   "20_TANKS_IP_DATA_RIO_04_FIRST_TANK_BWT_TEMP" : Real = PLC "20_TANKS_IP_DATA".RIO_04.FIRST_TANK.BWT_TEMP, 1 s
   "20_TANKS_IP_DATA_RIO_04_FIRST_TANK_BWT_DO" : Real = PLC "20_TANKS_IP_DATA".RIO_04.FIRST_TANK.BWT_DO, 1 s
   "20_TANKS_IP_DATA_RIO_04_FIRST_TANK_BWT_PH" : Real = PLC "20_TANKS_IP_DATA".RIO_04.FIRST_TANK.BWT_PH, 1 s
   "20_TANKS_IP_DATA_RIO_06_FIRST_TANK_BWT_TEMP" : Real = PLC "20_TANKS_IP_DATA".RIO_06.FIRST_TANK.BWT_TEMP, 1 s
   "20_TANKS_IP_DATA_RIO_04_FIRST_TANK_BWT_LEVEL" : Real = PLC "20_TANKS_IP_DATA".RIO_04.FIRST_TANK.BWT_LEVEL, 1 s
   "504_Tank Grouping_DB2020_Tank12 Min Time_ET" : Time = PLC "504_Tank Grouping_DB2020"."Tank12 Min Time".ET, 1 s
   "20_TANKS_IP_DATA_RIO_06_SECOND_TANK_BWT_LEVEL" : Real = PLC "20_TANKS_IP_DATA".RIO_06.SECOND_TANK.BWT_LEVEL, 1 s
   "504_Tank Grouping_DB2020_Time Left Tank_Time Left Tank 13" : Real = PLC "504_Tank Grouping_DB2020"."Time Left Tank"."Time Left Tank 13", 1 s
   "504_Tank Grouping_DB2020_Time Left Tank_Time Left Tank 12" : Real = PLC "504_Tank Grouping_DB2020"."Time Left Tank"."Time Left Tank 12", 1 s
   "504_Tank Grouping_DB2020_Time Left Tank_Time Left Tank 11" : Real = PLC "504_Tank Grouping_DB2020"."Time Left Tank"."Time Left Tank 11", 1 s
   "504_Tank Grouping_DB2020_Time Left Tank_Time Left Tank 10" : Real = PLC "504_Tank Grouping_DB2020"."Time Left Tank"."Time Left Tank 10", 1 s
   "504_Tank Grouping_DB2020_Time Left Tank_Time Left Tank 9" : Real = PLC "504_Tank Grouping_DB2020"."Time Left Tank"."Time Left Tank 9", 1 s
   "504_Tank Grouping_DB2020_Time Left Tank_Time Left Tank 8" : Real = PLC "504_Tank Grouping_DB2020"."Time Left Tank"."Time Left Tank 8", 1 s
   "504_Tank Grouping_DB2020_Time Left Tank_Time Left Tank 6" : Real = PLC "504_Tank Grouping_DB2020"."Time Left Tank"."Time Left Tank 6", 1 s
   "504_Tank Grouping_DB2020_Time Left Tank_Time Left Tank 5" : Real = PLC "504_Tank Grouping_DB2020"."Time Left Tank"."Time Left Tank 5", 1 s
   "504_Tank Grouping_DB2020_Time Left Tank_Time Left Tank 4" : Real = PLC "504_Tank Grouping_DB2020"."Time Left Tank"."Time Left Tank 4", 1 s
   "504_Tank Grouping_DB2020_Time Left Tank_Time Left Tank 3" : Real = PLC "504_Tank Grouping_DB2020"."Time Left Tank"."Time Left Tank 3", 1 s
   "504_Tank Grouping_DB2020_Time Left Tank_Time Left Tank 2" : Real = PLC "504_Tank Grouping_DB2020"."Time Left Tank"."Time Left Tank 2", 1 s
   "504_Tank Grouping_DB2020_Time Left Tank_Time Left Tank 7" : Real = PLC "504_Tank Grouping_DB2020"."Time Left Tank"."Time Left Tank 7", 1 s
   "504_Tank Grouping_DB2020_Offset Timer_ET" : Time = PLC "504_Tank Grouping_DB2020"."Offset Timer".ET, 1 s
   "80_From_HMI_Test Tank Request" : Bool = PLC "80_From_HMI"."Test Tank Request", 1 s
   "504_Tank Grouping_DB2020_RUN" : Bool = PLC "504_Tank Grouping_DB2020".RUN, 1 s
   "20_TANKS_IP_DATA_RIO_07_FIRST_TANK_BWT_TEMP" : Real = PLC "20_TANKS_IP_DATA".RIO_07.FIRST_TANK.BWT_TEMP, 1 s
   "20_TANKS_IP_DATA_RIO_07_FIRST_TANK_BWT_DO" : Real = PLC "20_TANKS_IP_DATA".RIO_07.FIRST_TANK.BWT_DO, 1 s
   "20_TANKS_IP_DATA_RIO_07_FIRST_TANK_BWT_PH" : Real = PLC "20_TANKS_IP_DATA".RIO_07.FIRST_TANK.BWT_PH, 1 s
   "20_TANKS_IP_DATA_RIO_07_FIRST_TANK_BWT_LEVEL" : Real = PLC "20_TANKS_IP_DATA".RIO_07.FIRST_TANK.BWT_LEVEL, 1 s
   "20_TANKS_IP_DATA_RIO_07_FIRST_TANK_TANKS_PRESS" : Real = PLC "20_TANKS_IP_DATA".RIO_07.FIRST_TANK.TANKS_PRESS, 1 s
   "504_Tank Grouping_DB2020_Tank14 Min Time_ET" : Time = PLC "504_Tank Grouping_DB2020"."Tank14 Min Time".ET, 1 s
   "504_Tank Grouping_DB2020_Tank13 Min Time_ET" : Time = PLC "504_Tank Grouping_DB2020"."Tank13 Min Time".ET, 1 s
   "20_TANKS_IP_DATA_RIO_06_SECOND_TANK_BWT_TEMP" : Real = PLC "20_TANKS_IP_DATA".RIO_06.SECOND_TANK.BWT_TEMP, 1 s
   "20_TANKS_IP_DATA_RIO_06_SECOND_TANK_BWT_DO" : Real = PLC "20_TANKS_IP_DATA".RIO_06.SECOND_TANK.BWT_DO, 1 s
   "20_TANKS_IP_DATA_RIO_06_SECOND_TANK_BWT_PH" : Real = PLC "20_TANKS_IP_DATA".RIO_06.SECOND_TANK.BWT_PH, 1 s
   "20_TANKS_IP_DATA_RIO_06_SECOND_TANK_TANKS_PRESS" : Real = PLC "20_TANKS_IP_DATA".RIO_06.SECOND_TANK.TANKS_PRESS, 1 s
   "20_TANKS_IP_DATA_RIO_04_FIRST_TANK_TANKS_PRESS" : Real = PLC "20_TANKS_IP_DATA".RIO_04.FIRST_TANK.TANKS_PRESS, 1 s
   "504_Tank Grouping_DB2020_Tank7 Min Time_ET" : Time = PLC "504_Tank Grouping_DB2020"."Tank7 Min Time".ET, 1 s
   "20_TANKS_IP_DATA_RIO_03_SECOND_TANK_BWT_TEMP" : Real = PLC "20_TANKS_IP_DATA".RIO_03.SECOND_TANK.BWT_TEMP, 1 s
   "504_Tank Grouping_DB2020_Sequence Time m Offset" : Time = PLC "504_Tank Grouping_DB2020"."Sequence Time m Offset", 1 s
   "504_Tank Grouping_DB2020_RUN TANK 13" : Bool = PLC "504_Tank Grouping_DB2020"."RUN TANK 13", 1 s
   "504_Tank Grouping_DB2020_RUN TANK 12" : Bool = PLC "504_Tank Grouping_DB2020"."RUN TANK 12", 1 s
   "504_Tank Grouping_DB2020_RUN TANK 11" : Bool = PLC "504_Tank Grouping_DB2020"."RUN TANK 11", 1 s
   "504_Tank Grouping_DB2020_RUN TANK 10" : Bool = PLC "504_Tank Grouping_DB2020"."RUN TANK 10", 1 s
   "504_Tank Grouping_DB2020_RUN TANK 9" : Bool = PLC "504_Tank Grouping_DB2020"."RUN TANK 9", 1 s
   "504_Tank Grouping_DB2020_RUN TANK 8" : Bool = PLC "504_Tank Grouping_DB2020"."RUN TANK 8", 1 s
   "504_Tank Grouping_DB2020_RUN TANK 6" : Bool = PLC "504_Tank Grouping_DB2020"."RUN TANK 6", 1 s
   "504_Tank Grouping_DB2020_RUN TANK 14" : Bool = PLC "504_Tank Grouping_DB2020"."RUN TANK 14", 1 s
   "20_TANKS_IP_DATA_RIO_07_FIRST_TANK_MBG_FLOW" : Real = PLC "20_TANKS_IP_DATA".RIO_07.FIRST_TANK.MBG_FLOW, 1 s
   "20_TANKS_IP_DATA_RIO_07_FIRST_TANK_USD_FLOW" : Real = PLC "20_TANKS_IP_DATA".RIO_07.FIRST_TANK.USD_FLOW, 1 s
   "20_TANKS_IP_DATA_RIO_07_FIRST_TANK_GTT_ISOL_VALVE_CLSD" : Bool = PLC "20_TANKS_IP_DATA".RIO_07.FIRST_TANK.GTT_ISOL_VALVE_CLSD, 1 s
   "20_TANKS_IP_DATA_RIO_07_FIRST_TANK_GTT_ISOL_VALVE_OPEN" : Bool = PLC "20_TANKS_IP_DATA".RIO_07.FIRST_TANK.GTT_ISOL_VALVE_OPEN, 1 s
   "20_TANKS_IP_DATA_RIO_07_FIRST_TANK_BWT_LEVEL_HIHI" : Bool = PLC "20_TANKS_IP_DATA".RIO_07.FIRST_TANK.BWT_LEVEL_HIHI, 1 s
   "20_TANKS_IP_DATA_RIO_06_SECOND_TANK_GTT_ISOL_VALVE_CLSD" : Bool = PLC "20_TANKS_IP_DATA".RIO_06.SECOND_TANK.GTT_ISOL_VALVE_CLSD, 1 s
   "20_TANKS_IP_DATA_RIO_06_SECOND_TANK_GTT_ISOL_VALVE_OPEN" : Bool = PLC "20_TANKS_IP_DATA".RIO_06.SECOND_TANK.GTT_ISOL_VALVE_OPEN, 1 s
   "Tank 3S BWT Level High High Switch" : Bool = PLC "Tank 3S BWT Level High High Switch" AT %I33.2, 1 s
   "20_TANKS_IP_DATA_RIO_06_SECOND_TANK_USD_FLOW" : Real = PLC "20_TANKS_IP_DATA".RIO_06.SECOND_TANK.USD_FLOW, 1 s
   "20_TANKS_IP_DATA_RIO_06_SECOND_TANK_BWT_LEVEL_HIHI" : Bool = PLC "20_TANKS_IP_DATA".RIO_06.SECOND_TANK.BWT_LEVEL_HIHI, 1 s
   "20_TANKS_IP_DATA_RIO_06_FIRST_TANK_GTT_ISOL_VALVE_CLSD" : Bool = PLC "20_TANKS_IP_DATA".RIO_06.FIRST_TANK.GTT_ISOL_VALVE_CLSD, 1 s
   "20_TANKS_IP_DATA_RIO_06_FIRST_TANK_GTT_ISOL_VALVE_OPEN" : Bool = PLC "20_TANKS_IP_DATA".RIO_06.FIRST_TANK.GTT_ISOL_VALVE_OPEN, 1 s
   "20_TANKS_IP_DATA_RIO_06_FIRST_TANK_MBG_FLOW" : Real = PLC "20_TANKS_IP_DATA".RIO_06.FIRST_TANK.MBG_FLOW, 1 s
   "20_TANKS_IP_DATA_RIO_06_FIRST_TANK_USD_FLOW" : Real = PLC "20_TANKS_IP_DATA".RIO_06.FIRST_TANK.USD_FLOW, 1 s
   "20_TANKS_IP_DATA_RIO_06_FIRST_TANK_BWT_LEVEL_HIHI" : Bool = PLC "20_TANKS_IP_DATA".RIO_06.FIRST_TANK.BWT_LEVEL_HIHI, 1 s
   "20_TANKS_IP_DATA_RIO_05_SECOND_TANK_GTT_ISOL_VALVE_CLSD" : Bool = PLC "20_TANKS_IP_DATA".RIO_05.SECOND_TANK.GTT_ISOL_VALVE_CLSD, 1 s
   "20_TANKS_IP_DATA_RIO_01_FIRST_TANK_TANKS_PRESS" : Real = PLC "20_TANKS_IP_DATA".RIO_01.FIRST_TANK.TANKS_PRESS, 1 s
   "20_TANKS_IP_DATA_RIO_01_FIRST_TANK_BWT_LEVEL" : Real = PLC "20_TANKS_IP_DATA".RIO_01.FIRST_TANK.BWT_LEVEL, 1 s
   "20_TANKS_IP_DATA_RIO_01_FIRST_TANK_BWT_PH" : Real = PLC "20_TANKS_IP_DATA".RIO_01.FIRST_TANK.BWT_PH, 1 s
   "20_TANKS_IP_DATA_RIO_01_FIRST_TANK_BWT_DO" : Real = PLC "20_TANKS_IP_DATA".RIO_01.FIRST_TANK.BWT_DO, 1 s
   "20_TANKS_IP_DATA_RIO_03_SECOND_TANK_BWT_DO" : Real = PLC "20_TANKS_IP_DATA".RIO_03.SECOND_TANK.BWT_DO, 1 s
   "20_TANKS_IP_DATA_RIO_03_SECOND_TANK_BWT_PH" : Real = PLC "20_TANKS_IP_DATA".RIO_03.SECOND_TANK.BWT_PH, 1 s
   "20_TANKS_IP_DATA_RIO_03_SECOND_TANK_BWT_LEVEL" : Real = PLC "20_TANKS_IP_DATA".RIO_03.SECOND_TANK.BWT_LEVEL, 1 s
   "20_TANKS_IP_DATA_RIO_03_SECOND_TANK_TANKS_PRESS" : Real = PLC "20_TANKS_IP_DATA".RIO_03.SECOND_TANK.TANKS_PRESS, 1 s
   "504_Tank Grouping_DB2020_Tank6 Min Time_ET" : Time = PLC "504_Tank Grouping_DB2020"."Tank6 Min Time".ET, 1 s
   "20_TANKS_IP_DATA_RIO_03_FIRST_TANK_BWT_TEMP" : Real = PLC "20_TANKS_IP_DATA".RIO_03.FIRST_TANK.BWT_TEMP, 1 s
   "20_TANKS_IP_DATA_RIO_03_FIRST_TANK_BWT_DO" : Real = PLC "20_TANKS_IP_DATA".RIO_03.FIRST_TANK.BWT_DO, 1 s
   "20_TANKS_IP_DATA_RIO_03_FIRST_TANK_BWT_PH" : Real = PLC "20_TANKS_IP_DATA".RIO_03.FIRST_TANK.BWT_PH, 1 s
   "20_TANKS_IP_DATA_RIO_03_FIRST_TANK_BWT_LEVEL" : Real = PLC "20_TANKS_IP_DATA".RIO_03.FIRST_TANK.BWT_LEVEL, 1 s
   "20_TANKS_IP_DATA_RIO_03_FIRST_TANK_TANKS_PRESS" : Real = PLC "20_TANKS_IP_DATA".RIO_03.FIRST_TANK.TANKS_PRESS, 1 s
   "504_Tank Grouping_DB2020_Tank5 Min Time_ET" : Time = PLC "504_Tank Grouping_DB2020"."Tank5 Min Time".ET, 1 s
   "504_Tank Grouping_DB2020_Tank3 Min Time_ET" : Time = PLC "504_Tank Grouping_DB2020"."Tank3 Min Time".ET, 1 s
   "20_TANKS_IP_DATA_RIO_05_SECOND_TANK_MBG_FLOW" : Real = PLC "20_TANKS_IP_DATA".RIO_05.SECOND_TANK.MBG_FLOW, 1 s
   "504_Tank Grouping_DB2020_Tank4 Min Time_ET" : Time = PLC "504_Tank Grouping_DB2020"."Tank4 Min Time".ET, 1 s
   "20_TANKS_IP_DATA_RIO_01_THIRD_TANK_BWT_DO" : Real = PLC "20_TANKS_IP_DATA".RIO_01.THIRD_TANK.BWT_DO, 1 s
   "20_TANKS_IP_DATA_RIO_01_THIRD_TANK_BWT_PH" : Real = PLC "20_TANKS_IP_DATA".RIO_01.THIRD_TANK.BWT_PH, 1 s
   "20_TANKS_IP_DATA_RIO_01_THIRD_TANK_BWT_LEVEL" : Real = PLC "20_TANKS_IP_DATA".RIO_01.THIRD_TANK.BWT_LEVEL, 1 s
   "20_TANKS_IP_DATA_RIO_01_THIRD_TANK_TANKS_PRESS" : Real = PLC "20_TANKS_IP_DATA".RIO_01.THIRD_TANK.TANKS_PRESS, 1 s
   "20_TANKS_IP_DATA_RIO_01_SECOND_TANK_BWT_TEMP" : Real = PLC "20_TANKS_IP_DATA".RIO_01.SECOND_TANK.BWT_TEMP, 1 s
   "20_TANKS_IP_DATA_RIO_01_SECOND_TANK_BWT_DO" : Real = PLC "20_TANKS_IP_DATA".RIO_01.SECOND_TANK.BWT_DO, 1 s
   "20_TANKS_IP_DATA_RIO_01_SECOND_TANK_BWT_PH" : Real = PLC "20_TANKS_IP_DATA".RIO_01.SECOND_TANK.BWT_PH, 1 s
   "20_TANKS_IP_DATA_RIO_01_SECOND_TANK_BWT_LEVEL" : Real = PLC "20_TANKS_IP_DATA".RIO_01.SECOND_TANK.BWT_LEVEL, 1 s
   "20_TANKS_IP_DATA_RIO_01_SECOND_TANK_TANKS_PRESS" : Real = PLC "20_TANKS_IP_DATA".RIO_01.SECOND_TANK.TANKS_PRESS, 1 s
   "504_Tank Grouping_DB2020_Tank2 Min Time_ET" : Time = PLC "504_Tank Grouping_DB2020"."Tank2 Min Time".ET, 1 s
   "504_Tank Grouping_DB2020_Tank1 Min Time_ET" : Time = PLC "504_Tank Grouping_DB2020"."Tank1 Min Time".ET, 1 s
   "20_TANKS_IP_DATA_RIO_01_FIRST_TANK_BWT_TEMP" : Real = PLC "20_TANKS_IP_DATA".RIO_01.FIRST_TANK.BWT_TEMP, 1 s
   "20_TANKS_IP_DATA_RIO_01_THIRD_TANK_BWT_TEMP" : Real = PLC "20_TANKS_IP_DATA".RIO_01.THIRD_TANK.BWT_TEMP, 1 s
   "RIO3_SPR_DI_33_3" : Bool = PLC RIO3_SPR_DI_33_3 AT %I33.3, 1 s
   "150_GCU_LCL_CNTRL_DB_LCL_CNTRL_ACTV" : Bool = PLC "150_GCU_LCL_CNTRL_DB".LCL_CNTRL_ACTV, 1 s
   "RIO3_SPR_DI_33_5" : Bool = PLC RIO3_SPR_DI_33_5 AT %I33.5, 1 s
   "TT426_5S_ALM_ANALOG_DB_VERY LOW LEVEL VALUE (LL)" : Real = PLC TT426_5S_ALM_ANALOG_DB."VERY LOW LEVEL VALUE (LL)" AT %DB2082.DBD22, 1 s
   "TT426_5S_ALM_ANALOG_DB_LOW LEVEL VALUE (L)" : Real = PLC TT426_5S_ALM_ANALOG_DB."LOW LEVEL VALUE (L)" AT %DB2082.DBD26, 1 s
   "TT426_5S_ALM_ANALOG_DB_HIGH LEVEL VALUE (H)" : Real = PLC TT426_5S_ALM_ANALOG_DB."HIGH LEVEL VALUE (H)" AT %DB2082.DBD30, 1 s
   "TT426_5S_ALM_ANALOG_DB_VERY HIGH LEVEL VALUE (HH)" : Real = PLC TT426_5S_ALM_ANALOG_DB."VERY HIGH LEVEL VALUE (HH)" AT %DB2082.DBD34, 1 s
   "TT426STR_ALM_ANALOG_DB_VERY LOW LEVEL VALUE (LL)" : Real = PLC TT426STR_ALM_ANALOG_DB."VERY LOW LEVEL VALUE (LL)" AT %DB2072.DBD22, 1 s
   "TT426STR_ALM_ANALOG_DB_LOW LEVEL VALUE (L)" : Real = PLC TT426STR_ALM_ANALOG_DB."LOW LEVEL VALUE (L)" AT %DB2072.DBD26, 1 s
   "TT426STR_ALM_ANALOG_DB_HIGH LEVEL VALUE (H)" : Real = PLC TT426STR_ALM_ANALOG_DB."HIGH LEVEL VALUE (H)" AT %DB2072.DBD30, 1 s
   "TT426STR_ALM_ANALOG_DB_VERY HIGH LEVEL VALUE (HH)" : Real = PLC TT426STR_ALM_ANALOG_DB."VERY HIGH LEVEL VALUE (HH)" AT %DB2072.DBD34, 1 s
   "TT426PORT_ALM_ANALOG_DB_VERY LOW LEVEL VALUE (LL)" : Real = PLC TT426PORT_ALM_ANALOG_DB."VERY LOW LEVEL VALUE (LL)" AT %DB2071.DBD22, 1 s
   "TT426PORT_ALM_ANALOG_DB_LOW LEVEL VALUE (L)" : Real = PLC TT426PORT_ALM_ANALOG_DB."LOW LEVEL VALUE (L)" AT %DB2071.DBD26, 1 s
   "TT426PORT_ALM_ANALOG_DB_HIGH LEVEL VALUE (H)" : Real = PLC TT426PORT_ALM_ANALOG_DB."HIGH LEVEL VALUE (H)" AT %DB2071.DBD30, 1 s
   "TT426PORT_ALM_ANALOG_DB_VERY HIGH LEVEL VALUE (HH)" : Real = PLC TT426PORT_ALM_ANALOG_DB."VERY HIGH LEVEL VALUE (HH)" AT %DB2071.DBD34, 1 s
   "PIT424PORT_ALM_ANALOG_DB_VERY HIGH LEVEL VALUE (HH)" : Real = PLC PIT424PORT_ALM_ANALOG_DB."VERY HIGH LEVEL VALUE (HH)" AT %DB2070.DBD34, 1 s
   "LIT304_ALM_ANALOG_DB71_VERY LOW LEVEL VALUE (LL)" : Real = PLC LIT304_ALM_ANALOG_DB71."VERY LOW LEVEL VALUE (LL)" AT %DB71.DBD22, 1 s
   "LIT304_ALM_ANALOG_DB71_LOW LEVEL VALUE (L)" : Real = PLC LIT304_ALM_ANALOG_DB71."LOW LEVEL VALUE (L)" AT %DB71.DBD26, 1 s
   "LIT304_ALM_ANALOG_DB71_HIGH LEVEL VALUE (H)" : Real = PLC LIT304_ALM_ANALOG_DB71."HIGH LEVEL VALUE (H)" AT %DB71.DBD30, 1 s
   "LIT304_ALM_ANALOG_DB71_VERY HIGH LEVEL VALUE (HH)" : Real = PLC LIT304_ALM_ANALOG_DB71."VERY HIGH LEVEL VALUE (HH)" AT %DB71.DBD34, 1 s
   "TIT406_ALM_ANALOG_DB74_VERY LOW LEVEL VALUE (LL)" : Real = PLC TIT406_ALM_ANALOG_DB74."VERY LOW LEVEL VALUE (LL)" AT %DB74.DBD22, 1 s
   "TIT406_ALM_ANALOG_DB74_LOW LEVEL VALUE (L)" : Real = PLC TIT406_ALM_ANALOG_DB74."LOW LEVEL VALUE (L)" AT %DB74.DBD26, 1 s
   "TIT406_ALM_ANALOG_DB74_HIGH LEVEL VALUE (H)" : Real = PLC TIT406_ALM_ANALOG_DB74."HIGH LEVEL VALUE (H)" AT %DB74.DBD30, 1 s
   "TIT406_ALM_ANALOG_DB74_VERY HIGH LEVEL VALUE (HH)" : Real = PLC TIT406_ALM_ANALOG_DB74."VERY HIGH LEVEL VALUE (HH)" AT %DB74.DBD34, 1 s
   "PIT424_RIO6_ALM_ANALOG_DB_VERY HIGH LEVEL VALUE (HH)" : Real = PLC PIT424_RIO6_ALM_ANALOG_DB."VERY HIGH LEVEL VALUE (HH)" AT %DB2223.DBD34, 1 s
   "PIT424_RIO6_ALM_ANALOG_DB_HIGH LEVEL VALUE (H)" : Real = PLC PIT424_RIO6_ALM_ANALOG_DB."HIGH LEVEL VALUE (H)" AT %DB2223.DBD30, 1 s
   "PIT424_RIO6_ALM_ANALOG_DB_LOW LEVEL VALUE (L)" : Real = PLC PIT424_RIO6_ALM_ANALOG_DB."LOW LEVEL VALUE (L)" AT %DB2223.DBD26, 1 s
   "PIT424_RIO6_ALM_ANALOG_DB_VERY LOW LEVEL VALUE (LL)" : Real = PLC PIT424_RIO6_ALM_ANALOG_DB."VERY LOW LEVEL VALUE (LL)" AT %DB2223.DBD22, 1 s
   "TT426_5P_ALM_ANALOG_DB_HIGH LEVEL VALUE (H)" : Real = PLC TT426_5P_ALM_ANALOG_DB."HIGH LEVEL VALUE (H)" AT %DB2081.DBD30, 1 s
   "TT426_5P_ALM_ANALOG_DB_VERY HIGH LEVEL VALUE (HH)" : Real = PLC TT426_5P_ALM_ANALOG_DB."VERY HIGH LEVEL VALUE (HH)" AT %DB2081.DBD34, 1 s
   "PIT424_RIO5_ALM_ANALOG_DB_VERY LOW LEVEL VALUE (LL)" : Real = PLC PIT424_RIO5_ALM_ANALOG_DB."VERY LOW LEVEL VALUE (LL)" AT %DB2222.DBD22, 1 s
   "PIT424_RIO5_ALM_ANALOG_DB_LOW LEVEL VALUE (L)" : Real = PLC PIT424_RIO5_ALM_ANALOG_DB."LOW LEVEL VALUE (L)" AT %DB2222.DBD26, 1 s
   "PIT424_RIO5_ALM_ANALOG_DB_HIGH LEVEL VALUE (H)" : Real = PLC PIT424_RIO5_ALM_ANALOG_DB."HIGH LEVEL VALUE (H)" AT %DB2222.DBD30, 1 s
   "PIT424_RIO5_ALM_ANALOG_DB_VERY HIGH LEVEL VALUE (HH)" : Real = PLC PIT424_RIO5_ALM_ANALOG_DB."VERY HIGH LEVEL VALUE (HH)" AT %DB2222.DBD34, 1 s
   "TT426_APT_ALM_ANALOG_DB_VERY LOW LEVEL VALUE (LL)" : Real = PLC TT426_APT_ALM_ANALOG_DB."VERY LOW LEVEL VALUE (LL)" AT %DB2087.DBD22, 1 s
   "TT426_APT_ALM_ANALOG_DB_LOW LEVEL VALUE (L)" : Real = PLC TT426_APT_ALM_ANALOG_DB."LOW LEVEL VALUE (L)" AT %DB2087.DBD26, 1 s
   "TT426_APT_ALM_ANALOG_DB_HIGH LEVEL VALUE (H)" : Real = PLC TT426_APT_ALM_ANALOG_DB."HIGH LEVEL VALUE (H)" AT %DB2087.DBD30, 1 s
   "TT426_APT_ALM_ANALOG_DB_VERY HIGH LEVEL VALUE (HH)" : Real = PLC TT426_APT_ALM_ANALOG_DB."VERY HIGH LEVEL VALUE (HH)" AT %DB2087.DBD34, 1 s
   "502_ALM_ANALOG_IDB PIT 416_VERY LOW LEVEL VALUE (LL)" : Real = PLC "502_ALM_ANALOG_IDB PIT 416"."VERY LOW LEVEL VALUE (LL)" AT %DB65.DBD22, 1 s
   "PIT424_RIO7_ALM_ANALOG_DB_VERY LOW LEVEL VALUE (LL)" : Real = PLC PIT424_RIO7_ALM_ANALOG_DB."VERY LOW LEVEL VALUE (LL)" AT %DB2224.DBD22, 1 s
   "PIT424_RIO7_ALM_ANALOG_DB_HIGH LEVEL VALUE (H)" : Real = PLC PIT424_RIO7_ALM_ANALOG_DB."HIGH LEVEL VALUE (H)" AT %DB2224.DBD30, 1 s
   "PIT424_RIO7_ALM_ANALOG_DB_VERY HIGH LEVEL VALUE (HH)" : Real = PLC PIT424_RIO7_ALM_ANALOG_DB."VERY HIGH LEVEL VALUE (HH)" AT %DB2224.DBD34, 1 s
   "TT426_6S_ALM_ANALOG_DB_VERY LOW LEVEL VALUE (LL)" : Real = PLC TT426_6S_ALM_ANALOG_DB."VERY LOW LEVEL VALUE (LL)" AT %DB2085.DBD22, 1 s
   "TT426_6S_ALM_ANALOG_DB_LOW LEVEL VALUE (L)" : Real = PLC TT426_6S_ALM_ANALOG_DB."LOW LEVEL VALUE (L)" AT %DB2085.DBD26, 1 s
   "TT426_6S_ALM_ANALOG_DB_HIGH LEVEL VALUE (H)" : Real = PLC TT426_6S_ALM_ANALOG_DB."HIGH LEVEL VALUE (H)" AT %DB2085.DBD30, 1 s
   "TT426_6S_ALM_ANALOG_DB_VERY HIGH LEVEL VALUE (HH)" : Real = PLC TT426_6S_ALM_ANALOG_DB."VERY HIGH LEVEL VALUE (HH)" AT %DB2085.DBD34, 1 s
   "TT426_6P_ALM_ANALOG_DB_VERY LOW LEVEL VALUE (LL)" : Real = PLC TT426_6P_ALM_ANALOG_DB."VERY LOW LEVEL VALUE (LL)" AT %DB2083.DBD22, 1 s
   "TT426_6P_ALM_ANALOG_DB_LOW LEVEL VALUE (L)" : Real = PLC TT426_6P_ALM_ANALOG_DB."LOW LEVEL VALUE (L)" AT %DB2083.DBD26, 1 s
   "TT426_6P_ALM_ANALOG_DB_HIGH LEVEL VALUE (H)" : Real = PLC TT426_6P_ALM_ANALOG_DB."HIGH LEVEL VALUE (H)" AT %DB2083.DBD30, 1 s
   "TT426_6P_ALM_ANALOG_DB_VERY HIGH LEVEL VALUE (HH)" : Real = PLC TT426_6P_ALM_ANALOG_DB."VERY HIGH LEVEL VALUE (HH)" AT %DB2083.DBD34, 1 s
   "PIT424_RIO7_ALM_ANALOG_DB_LOW LEVEL VALUE (L)" : Real = PLC PIT424_RIO7_ALM_ANALOG_DB."LOW LEVEL VALUE (L)" AT %DB2224.DBD26, 1 s
   "502_ALM_ANALOG_IDB PIT 416_LOW LEVEL VALUE (L)" : Real = PLC "Sequence Times_DB"."Treatment Timer"."Minutes Left" AT %DB65.DBD26, 1 s
   "502_ALM_ANALOG_IDB PIT 416_HIGH LEVEL VALUE (H)" : Real = PLC "502_ALM_ANALOG_IDB PIT 416"."HIGH LEVEL VALUE (H)" AT %DB65.DBD30, 1 s
   "502_ALM_ANALOG_IDB PIT 416_VERY HIGH LEVEL VALUE (HH)" : Real = PLC "502_ALM_ANALOG_IDB PIT 416"."VERY HIGH LEVEL VALUE (HH)" AT %DB65.DBD34, 1 s
   "PT415_RIO4_ALM_ANALOG_DB_HIGH LEVEL VALUE (H)" : Real = PLC PT415_RIO4_ALM_ANALOG_DB."HIGH LEVEL VALUE (H)" AT %DB2216.DBD30, 1 s
   "PT415_RIO4_ALM_ANALOG_DB_VERY HIGH LEVEL VALUE (HH)" : Real = PLC PT415_RIO4_ALM_ANALOG_DB."VERY HIGH LEVEL VALUE (HH)" AT %DB2216.DBD34, 1 s
   "TT426_FPT_ALM_ANALOG_DB_VERY LOW LEVEL VALUE (LL)" : Real = PLC TT426_FPT_ALM_ANALOG_DB."VERY LOW LEVEL VALUE (LL)" AT %DB2074.DBD22, 1 s
   "TT426_FPT_ALM_ANALOG_DB_LOW LEVEL VALUE (L)" : Real = PLC TT426_FPT_ALM_ANALOG_DB."LOW LEVEL VALUE (L)" AT %DB2074.DBD26, 1 s
   "TT426_FPT_ALM_ANALOG_DB_HIGH LEVEL VALUE (H)" : Real = PLC TT426_FPT_ALM_ANALOG_DB."HIGH LEVEL VALUE (H)" AT %DB2074.DBD30, 1 s
   "TT426_FPT_ALM_ANALOG_DB_VERY HIGH LEVEL VALUE (HH)" : Real = PLC TT426_FPT_ALM_ANALOG_DB."VERY HIGH LEVEL VALUE (HH)" AT %DB2074.DBD34, 1 s
   "PIT424_RIO4_ALM_ANALOG_DB_VERY LOW LEVEL VALUE (LL)" : Real = PLC PIT424_RIO4_ALM_ANALOG_DB."VERY LOW LEVEL VALUE (LL)" AT %DB2221.DBD22, 1 s
   "PIT424_RIO4_ALM_ANALOG_DB_LOW LEVEL VALUE (L)" : Real = PLC PIT424_RIO4_ALM_ANALOG_DB."LOW LEVEL VALUE (L)" AT %DB2221.DBD26, 1 s
   "PIT424_RIO4_ALM_ANALOG_DB_HIGH LEVEL VALUE (H)" : Real = PLC PIT424_RIO4_ALM_ANALOG_DB."HIGH LEVEL VALUE (H)" AT %DB2221.DBD30, 1 s
   "PIT424_RIO4_ALM_ANALOG_DB_VERY HIGH LEVEL VALUE (HH)" : Real = PLC PIT424_RIO4_ALM_ANALOG_DB."VERY HIGH LEVEL VALUE (HH)" AT %DB2221.DBD34, 1 s
   "PT415_RIO4_ALM_ANALOG_DB_LOW LEVEL VALUE (L)" : Real = PLC PT415_RIO4_ALM_ANALOG_DB."LOW LEVEL VALUE (L)" AT %DB2216.DBD26, 1 s
   "TT426_3S_ALM_ANALOG_DB_VERY LOW LEVEL VALUE (LL)" : Real = PLC TT426_3S_ALM_ANALOG_DB."VERY LOW LEVEL VALUE (LL)" AT %DB2078.DBD22, 1 s
   "TT426_3S_ALM_ANALOG_DB_HIGH LEVEL VALUE (H)" : Real = PLC TT426_3S_ALM_ANALOG_DB."HIGH LEVEL VALUE (H)" AT %DB2078.DBD30, 1 s
   "TT426_3S_ALM_ANALOG_DB_VERY HIGH LEVEL VALUE (HH)" : Real = PLC TT426_3S_ALM_ANALOG_DB."VERY HIGH LEVEL VALUE (HH)" AT %DB2078.DBD34, 1 s
   "PIT424_RIO3_ALM_ANALOG_DB_VERY LOW LEVEL VALUE (LL)" : Real = PLC PIT424_RIO3_ALM_ANALOG_DB."VERY LOW LEVEL VALUE (LL)" AT %DB2220.DBD22, 1 s
   "PIT424_RIO3_ALM_ANALOG_DB_LOW LEVEL VALUE (L)" : Real = PLC PIT424_RIO3_ALM_ANALOG_DB."LOW LEVEL VALUE (L)" AT %DB2220.DBD26, 1 s
   "PIT424_RIO3_ALM_ANALOG_DB_HIGH LEVEL VALUE (H)" : Real = PLC PIT424_RIO3_ALM_ANALOG_DB."HIGH LEVEL VALUE (H)" AT %DB2220.DBD30, 1 s
   "PIT424_RIO3_ALM_ANALOG_DB_VERY HIGH LEVEL VALUE (HH)" : Real = PLC PIT424_RIO3_ALM_ANALOG_DB."VERY HIGH LEVEL VALUE (HH)" AT %DB2220.DBD34, 1 s
   "TT426_3P_ALM_ANALOG_DB_VERY LOW LEVEL VALUE (LL)" : Real = PLC TT426_3P_ALM_ANALOG_DB."VERY LOW LEVEL VALUE (LL)" AT %DB2077.DBD22, 1 s
   "TT426_3P_ALM_ANALOG_DB_LOW LEVEL VALUE (L)" : Real = PLC TT426_3P_ALM_ANALOG_DB."LOW LEVEL VALUE (L)" AT %DB2077.DBD26, 1 s
   "TT426_3P_ALM_ANALOG_DB_HIGH LEVEL VALUE (H)" : Real = PLC TT426_3P_ALM_ANALOG_DB."HIGH LEVEL VALUE (H)" AT %DB2077.DBD30, 1 s
   "TT426_3P_ALM_ANALOG_DB_VERY HIGH LEVEL VALUE (HH)" : Real = PLC TT426_3P_ALM_ANALOG_DB."VERY HIGH LEVEL VALUE (HH)" AT %DB2077.DBD34, 1 s
   "TT426_3S_ALM_ANALOG_DB_LOW LEVEL VALUE (L)" : Real = PLC TT426_3S_ALM_ANALOG_DB."LOW LEVEL VALUE (L)" AT %DB2078.DBD26, 1 s
   "TT426_5P_ALM_ANALOG_DB_LOW LEVEL VALUE (L)" : Real = PLC TT426_5P_ALM_ANALOG_DB."LOW LEVEL VALUE (L)" AT %DB2081.DBD26, 1 s
   "PT415_RIO4_ALM_ANALOG_DB_VERY LOW LEVEL VALUE (LL)" : Real = PLC PT415_RIO4_ALM_ANALOG_DB."VERY LOW LEVEL VALUE (LL)" AT %DB2216.DBD22, 1 s
   "PIT353_ALM_ANALOG_DB72_HIGH LEVEL VALUE (H)" : Real = PLC PIT353_ALM_ANALOG_DB72."HIGH LEVEL VALUE (H)" AT %DB72.DBD30, 1 s
   "PT415PORT_ALM_ANALOG_DB_VERY LOW LEVEL VALUE (LL)" : Real = PLC PT415PORT_ALM_ANALOG_DB."VERY LOW LEVEL VALUE (LL)" AT %DB2069.DBD22, 1 s
   "PT415PORT_ALM_ANALOG_DB_LOW LEVEL VALUE (L)" : Real = PLC PT415PORT_ALM_ANALOG_DB."LOW LEVEL VALUE (L)" AT %DB2069.DBD26, 1 s
   "PT415PORT_ALM_ANALOG_DB_HIGH LEVEL VALUE (H)" : Real = PLC PT415PORT_ALM_ANALOG_DB."HIGH LEVEL VALUE (H)" AT %DB2069.DBD30, 1 s
   "PT415PORT_ALM_ANALOG_DB_VERY HIGH LEVEL VALUE (HH)" : Real = PLC PT415PORT_ALM_ANALOG_DB."VERY HIGH LEVEL VALUE (HH)" AT %DB2069.DBD34, 1 s
   "TT002_ALM_ANALOG_DB76_VERY LOW LEVEL VALUE (LL)" : Real = PLC TT002_ALM_ANALOG_DB76."VERY LOW LEVEL VALUE (LL)" AT %DB76.DBD22, 1 s
   "TT002_ALM_ANALOG_DB76_LOW LEVEL VALUE (L)" : Real = PLC TT002_ALM_ANALOG_DB76."LOW LEVEL VALUE (L)" AT %DB76.DBD26, 1 s
   "TT002_ALM_ANALOG_DB76_HIGH LEVEL VALUE (H)" : Real = PLC TT002_ALM_ANALOG_DB76."HIGH LEVEL VALUE (H)" AT %DB76.DBD30, 1 s
   "TT002_ALM_ANALOG_DB76_VERY HIGH LEVEL VALUE (HH)" : Real = PLC TT002_ALM_ANALOG_DB76."VERY HIGH LEVEL VALUE (HH)" AT %DB76.DBD34, 1 s
   "PIT358_ALM_ANALOG_DB78_VERY LOW LEVEL VALUE (LL)" : Real = PLC PIT358_ALM_ANALOG_DB78."VERY LOW LEVEL VALUE (LL)" AT %DB78.DBD22, 1 s
   "PIT358_ALM_ANALOG_DB78_LOW LEVEL VALUE (L)" : Real = PLC PIT358_ALM_ANALOG_DB78."LOW LEVEL VALUE (L)" AT %DB78.DBD26, 1 s
   "PIT353_ALM_ANALOG_DB72_VERY HIGH LEVEL VALUE (HH)" : Real = PLC PIT353_ALM_ANALOG_DB72."VERY HIGH LEVEL VALUE (HH)" AT %DB72.DBD34, 1 s
   "PIT358_ALM_ANALOG_DB78_HIGH LEVEL VALUE (H)" : Real = PLC PIT358_ALM_ANALOG_DB78."HIGH LEVEL VALUE (H)" AT %DB78.DBD30, 1 s
   "PIT348_ALM_ANALOG_DB73_VERY LOW LEVEL VALUE (LL)" : Real = PLC PIT348_ALM_ANALOG_DB73."VERY LOW LEVEL VALUE (LL)" AT %DB73.DBD22, 1 s
   "PIT348_ALM_ANALOG_DB73_LOW LEVEL VALUE (L)" : Real = PLC PIT348_ALM_ANALOG_DB73."LOW LEVEL VALUE (L)" AT %DB73.DBD26, 1 s
   "PIT348_ALM_ANALOG_DB73_HIGH LEVEL VALUE (H)" : Real = PLC PIT348_ALM_ANALOG_DB73."HIGH LEVEL VALUE (H)" AT %DB73.DBD30, 1 s
   "PIT348_ALM_ANALOG_DB73_VERY HIGH LEVEL VALUE (HH)" : Real = PLC PIT348_ALM_ANALOG_DB73."VERY HIGH LEVEL VALUE (HH)" AT %DB73.DBD34, 1 s
   "TIT408_ALM_ANALOG_DB75_VERY LOW LEVEL VALUE (LL)" : Real = PLC TIT408_ALM_ANALOG_DB75."VERY LOW LEVEL VALUE (LL)" AT %DB75.DBD22, 1 s
   "TIT408_ALM_ANALOG_DB75_LOW LEVEL VALUE (L)" : Real = PLC TIT408_ALM_ANALOG_DB75."LOW LEVEL VALUE (L)" AT %DB75.DBD26, 1 s
   "TIT408_ALM_ANALOG_DB75_HIGH LEVEL VALUE (H)" : Real = PLC TIT408_ALM_ANALOG_DB75."HIGH LEVEL VALUE (H)" AT %DB75.DBD30, 1 s
   "TIT408_ALM_ANALOG_DB75_VERY HIGH LEVEL VALUE (HH)" : Real = PLC TIT408_ALM_ANALOG_DB75."VERY HIGH LEVEL VALUE (HH)" AT %DB75.DBD34, 1 s
   "PIT353_ALM_ANALOG_DB72_VERY LOW LEVEL VALUE (LL)" : Real = PLC PIT353_ALM_ANALOG_DB72."VERY LOW LEVEL VALUE (LL)" AT %DB72.DBD22, 1 s
   "PIT353_ALM_ANALOG_DB72_LOW LEVEL VALUE (L)" : Real = PLC PIT353_ALM_ANALOG_DB72."LOW LEVEL VALUE (L)" AT %DB72.DBD26, 1 s
   "PIT358_ALM_ANALOG_DB78_VERY HIGH LEVEL VALUE (HH)" : Real = PLC PIT358_ALM_ANALOG_DB78."VERY HIGH LEVEL VALUE (HH)" AT %DB78.DBD34, 1 s
   "TT426_1S_ALM_ANALOG_DB_VERY LOW LEVEL VALUE (LL)" : Real = PLC TT426_1S_ALM_ANALOG_DB."VERY LOW LEVEL VALUE (LL)" AT %DB2076.DBD22, 1 s
   "TT426_5P_ALM_ANALOG_DB_VERY LOW LEVEL VALUE (LL)" : Real = PLC TT426_5P_ALM_ANALOG_DB."VERY LOW LEVEL VALUE (LL)" AT %DB2081.DBD22, 1 s
   "TT426_4S_ALM_ANALOG_DB_HIGH LEVEL VALUE (H)" : Real = PLC TT426_4S_ALM_ANALOG_DB."HIGH LEVEL VALUE (H)" AT %DB2080.DBD30, 1 s
   "Sequence Times_DB_Re-Ox Timer_PT_HOURS" : Real = PLC "Sequence Times_DB"."Re-Ox Timer".PT_HOURS, 1 s
   "Sequence Times_DB_Re-Ox Timer_Days Left" : DInt = PLC "Sequence Times_DB"."Re-Ox Timer"."Days Left", 1 s
   "Sequence Times_DB_Re-Ox Timer_Hours Left" : DInt = PLC "Sequence Times_DB"."Re-Ox Timer"."Hours Left", 1 s
   "Sequence Times_DB_Re-Ox Timer_Minutes Left" : DInt = PLC "Sequence Times_DB"."Re-Ox Timer"."Minutes Left", 1 s
   "Sequence Times_DB_De-Ox Timer_Days Left" : DInt = PLC "Sequence Times_DB"."De-Ox Timer"."Days Left", 1 s
   "Sequence Times_DB_De-Ox Timer_Hours Left" : DInt = PLC "Sequence Times_DB"."De-Ox Timer"."Hours Left", 1 s
   "Sequence Times_DB_De-Ox Timer_Minutes Left" : DInt = PLC "Sequence Times_DB"."De-Ox Timer"."Minutes Left", 1 s
   "Sequence Times_DB_Dwell Timer_PT_HOURS" : Real = PLC "Sequence Times_DB"."Dwell Timer".PT_HOURS, 1 s
   "Sequence Times_DB_De-Ox Timer_PT_HOURS" : Real = PLC "Sequence Times_DB"."De-Ox Timer".PT_HOURS, 1 s
   "Sequence Times_DB_Dwell Timer_Days Left" : DInt = PLC "Sequence Times_DB"."Dwell Timer"."Days Left", 1 s
   "Sequence Times_DB_Dwell Timer_Hours Left" : DInt = PLC "Sequence Times_DB"."Dwell Timer"."Hours Left", 1 s
   "Sequence Times_DB_Dwell Timer_Minutes Left" : DInt = PLC "Sequence Times_DB"."Dwell Timer"."Minutes Left", 1 s
   "504_Tank Grouping_DB2020_O2 De-Ox Setpoint" : Real = PLC "504_Tank Grouping_DB2020"."O2 De-Ox Setpoint", 1 s
   "Sequence Times_DB_Treatment Timer_Days Left" : DInt = PLC "Sequence Times_DB"."Treatment Timer"."Days Left", 1 s
   "Sequence Times_DB_Treatment Timer_Hours Left" : DInt = PLC "Sequence Times_DB"."Treatment Timer"."Hours Left", 1 s
   "Sequence Times_DB_Treatment Timer_Minutes Left" : DInt = PLC "Sequence Times_DB"."Treatment Timer"."Minutes Left", 1 s
   "Sequence Times_DB_Pre-Dwell Timer_PT_HOURS" : Real = PLC "Sequence Times_DB"."Pre-Dwell Timer".PT_HOURS, 1 s
   "Sequence Times_DB_Treatment Timer_Days" : DInt = PLC "Sequence Times_DB"."Treatment Timer".Days, 1 s
   "Sequence Times_DB_Treatment Timer_Hours" : DInt = PLC "Sequence Times_DB"."Treatment Timer".Hours, 1 s
   "Sequence Times_DB_Treatment Timer_Minutes" : DInt = PLC "Sequence Times_DB"."Treatment Timer".Minutes, 1 s
   "Sequence Times_DB_Jurney Time" : Real = PLC "Sequence Times_DB"."Jurney Time", 1 s
   "Sequence Times_DB_Post-Dwell Timer_Minutes Left" : DInt = PLC "Sequence Times_DB"."Post-Dwell Timer"."Minutes Left", 1 s
   "Sequence Times_DB_Post-Dwell Timer_Hours Left" : DInt = PLC "Sequence Times_DB"."Post-Dwell Timer"."Hours Left", 1 s
   "Sequence Times_DB_Post-Dwell Timer_Days Left" : DInt = PLC "Sequence Times_DB"."Post-Dwell Timer"."Days Left", 1 s
   "Sequence Times_DB_Post-Dwell Timer_PT_HOURS" : Real = PLC "Sequence Times_DB"."Post-Dwell Timer".PT_HOURS, 1 s
   "Sequence Times_DB_Treatment Timer_Enable" : Bool = PLC "Sequence Times_DB"."Treatment Timer".Enable, 1 s
   "2086_Times_CV422_FPT_MAX_TRVL_TIME" : Time = PLC "2086_Times".CV422_FPT_MAX_TRVL_TIME, 1 s
   "2086_Times_CV422_1P_MAX_TRVL_TIME" : Time = PLC "2086_Times".CV422_1P_MAX_TRVL_TIME, 1 s
   "2086_Times_CV421_1S_MAX_TRVL_TIME" : Time = PLC "2086_Times".CV421_1S_MAX_TRVL_TIME, 1 s
   "2086_Times_CV422_2P_MAX_TRVL_TIME" : Time = PLC "2086_Times".CV422_2P_MAX_TRVL_TIME, 1 s
   "2086_Times_CV421_2S_MAX_TRVL_TIME" : Time = PLC "2086_Times".CV421_2S_MAX_TRVL_TIME, 1 s
   "2086_Times_CV422_3P_MAX_TRVL_TIME" : Time = PLC "2086_Times".CV422_3P_MAX_TRVL_TIME, 1 s
   "2086_Times_CV421_3S_MAX_TRVL_TIME" : Time = PLC "2086_Times".CV421_3S_MAX_TRVL_TIME, 1 s
   "2086_Times_CV422_4P_MAX_TRVL_TIME" : Time = PLC "2086_Times".CV422_4P_MAX_TRVL_TIME, 1 s
   "2086_Times_CV421_4S_MAX_TRVL_TIME" : Time = PLC "2086_Times".CV421_4S_MAX_TRVL_TIME, 1 s
   "Sequence Times_DB_Jurney Time FB_Hours Left" : Int = PLC "Sequence Times_DB"."Jurney Time FB"."Hours Left", 1 s
   "2086_Times_CV422_5P_MAX_TRVL_TIME" : Time = PLC "2086_Times".CV422_5P_MAX_TRVL_TIME, 1 s
   "2086_Times_CV421_6S_MAX_TRVL_TIME" : Time = PLC "2086_Times".CV421_6S_MAX_TRVL_TIME, 1 s
   "2086_Times_CV422_6P_MAX_TRVL_TIME" : Time = PLC "2086_Times".CV422_6P_MAX_TRVL_TIME, 1 s
   "2086_Times_CV422_APT_MAX_TRVL_TIME" : Time = PLC "2086_Times".CV422_APT_MAX_TRVL_TIME, 1 s
   "2068_Sys_Status_Data_Not BWT mode Warning" : Bool = PLC "2068_Sys_Status_Data"."Not BWT mode Warning" AT %DB1.DBX0.0, 1 s
      on ChangeValue: "BWT_Warning"()
   "Sequence Times_DB_De-Ox Time" : Real = PLC "Sequence Times_DB"."De-Ox Time", 1 s
   "Sequence Times_DB_De-Ox SP Time" : Real = PLC "Sequence Times_DB"."De-Ox SP Time", 1 s
   "Sequence Times_DB_Dwell Time" : Real = PLC "Sequence Times_DB"."Dwell Time", 1 s
   "Sequence Times_DB_Post-Dwell Time" : Real = PLC "Sequence Times_DB"."Post-Dwell Time", 1 s
   "Sequence Times_DB_Re-Ox Time" : Real = PLC "Sequence Times_DB"."Re-Ox Time", 1 s
   "Sequence Times_DB_Pre-Dwell Time" : Real = PLC "Sequence Times_DB"."Pre-Dwell Time", 1 s
   "2086_Times_CV421_5S_MAX_TRVL_TIME" : Time = PLC "2086_Times".CV421_5S_MAX_TRVL_TIME, 1 s
   "Sequence Times_DB_Jurney Time FB_Days Left" : Int = PLC "Sequence Times_DB"."Jurney Time FB"."Days Left", 1 s
   "Sequence Times_DB_Pre-Dwell Timer_Hours Left" : DInt = PLC "Sequence Times_DB"."Pre-Dwell Timer"."Hours Left", 1 s
   "Sequence Times_DB_Pre-Dwell Timer_Minutes Left" : DInt = PLC "Sequence Times_DB"."Pre-Dwell Timer"."Minutes Left", 1 s
   "PT415_RIO7_ALM_ANALOG_DB_VERY HIGH LEVEL VALUE (HH)" : Real = PLC PT415_RIO7_ALM_ANALOG_DB."VERY HIGH LEVEL VALUE (HH)" AT %DB2225.DBD34, 1 s
   "FIT418_2P_ALM_ANALOG_DB_VERY LOW LEVEL VALUE (LL)" : Real = PLC FIT418_2P_ALM_ANALOG_DB."VERY LOW LEVEL VALUE (LL)" AT %DB2064.DBD22, 1 s
   "FIT418_2P_ALM_ANALOG_DB_LOW LEVEL VALUE (L)" : Real = PLC FIT418_2P_ALM_ANALOG_DB."LOW LEVEL VALUE (L)" AT %DB2064.DBD26, 1 s
   "FIT418_2P_ALM_ANALOG_DB_HIGH LEVEL VALUE (H)" : Real = PLC FIT418_2P_ALM_ANALOG_DB."HIGH LEVEL VALUE (H)" AT %DB2064.DBD30, 1 s
   "FIT418_2P_ALM_ANALOG_DB_VERY HIGH LEVEL VALUE (HH)" : Real = PLC FIT418_2P_ALM_ANALOG_DB."VERY HIGH LEVEL VALUE (HH)" AT %DB2064.DBD34, 1 s
   "FIT420PORT_ALM_ANALOG_DB_VERY LOW LEVEL VALUE (LL)" : Real = PLC FIT420PORT_ALM_ANALOG_DB."VERY LOW LEVEL VALUE (LL)" AT %DB2065.DBD22, 1 s
   "FIT420PORT_ALM_ANALOG_DB_LOW LEVEL VALUE (L)" : Real = PLC FIT420PORT_ALM_ANALOG_DB."LOW LEVEL VALUE (L)" AT %DB2065.DBD26, 1 s
   "FIT420PORT_ALM_ANALOG_DB_HIGH LEVEL VALUE (H)" : Real = PLC FIT420PORT_ALM_ANALOG_DB."HIGH LEVEL VALUE (H)" AT %DB2065.DBD30, 1 s
   "FIT420PORT_ALM_ANALOG_DB_VERY HIGH LEVEL VALUE (HH)" : Real = PLC FIT420PORT_ALM_ANALOG_DB."VERY HIGH LEVEL VALUE (HH)" AT %DB2065.DBD34, 1 s
   "PIT424PORT_ALM_ANALOG_DB_VERY LOW LEVEL VALUE (LL)" : Real = PLC PIT424PORT_ALM_ANALOG_DB."VERY LOW LEVEL VALUE (LL)" AT %DB2070.DBD22, 1 s
   "PT415_RIO7_ALM_ANALOG_DB_HIGH LEVEL VALUE (H)" : Real = PLC PT415_RIO7_ALM_ANALOG_DB."HIGH LEVEL VALUE (H)" AT %DB2225.DBD30, 1 s
   "PIT424PORT_ALM_ANALOG_DB_LOW LEVEL VALUE (L)" : Real = PLC PIT424PORT_ALM_ANALOG_DB."LOW LEVEL VALUE (L)" AT %DB2070.DBD26, 1 s
   "FIT417_2S_ALM_ANALOG_DB_VERY LOW LEVEL VALUE (LL)" : Real = PLC FIT417_2S_ALM_ANALOG_DB."VERY LOW LEVEL VALUE (LL)" AT %DB2066.DBD22, 1 s
   "FIT417_2S_ALM_ANALOG_DB_LOW LEVEL VALUE (L)" : Real = PLC FIT417_2S_ALM_ANALOG_DB."LOW LEVEL VALUE (L)" AT %DB2066.DBD26, 1 s
   "FIT417_2S_ALM_ANALOG_DB_HIGH LEVEL VALUE (H)" : Real = PLC FIT417_2S_ALM_ANALOG_DB."HIGH LEVEL VALUE (H)" AT %DB2066.DBD30, 1 s
   "FIT417_2S_ALM_ANALOG_DB_VERY HIGH LEVEL VALUE (HH)" : Real = PLC FIT417_2S_ALM_ANALOG_DB."VERY HIGH LEVEL VALUE (HH)" AT %DB2066.DBD34, 1 s
   "FIT419_ALM_ANALOG_DB_VERY LOW LEVEL VALUE (LL)" : Real = PLC FIT419_ALM_ANALOG_DB."VERY LOW LEVEL VALUE (LL)" AT %DB2067.DBD22, 1 s
   "FIT419_ALM_ANALOG_DB_LOW LEVEL VALUE (L)" : Real = PLC FIT419_ALM_ANALOG_DB."LOW LEVEL VALUE (L)" AT %DB2067.DBD26, 1 s
   "FIT419_ALM_ANALOG_DB_HIGH LEVEL VALUE (H)" : Real = PLC FIT419_ALM_ANALOG_DB."HIGH LEVEL VALUE (H)" AT %DB2067.DBD30, 1 s
   "FIT419_ALM_ANALOG_DB_VERY HIGH LEVEL VALUE (HH)" : Real = PLC FIT419_ALM_ANALOG_DB."VERY HIGH LEVEL VALUE (HH)" AT %DB2067.DBD34, 1 s
   "TT426_4S_ALM_ANALOG_DB_VERY LOW LEVEL VALUE (LL)" : Real = PLC TT426_4S_ALM_ANALOG_DB."VERY LOW LEVEL VALUE (LL)" AT %DB2080.DBD22, 1 s